   Circle "Kreis_157" at 637,438 size 15x15
      Appearance <- "DB_SDC_ERRORS.EMS[XXX].FC_HOIST_2"
   Circle "Kreis_158" at 637,454 size 15x15
      Appearance <- "DB_SDC_ERRORS.EMS[XXX].FC_HOIST_2"
   Circle "Kreis_159" at 637,470 size 15x15
      Appearance <- "DB_SDC_ERRORS.EMS[XXX].FC_HOIST_2"
   Circle "Kreis_160" at 637,486 size 15x15
      Appearance <- "DB_SDC_ERRORS.EMS[XXX].FC_HOIST_2"
   TextField "Textfeld_248" at 1003,235 size 31x132; Text '501 502 503 504 505 506 507 508 Command forward 501'
   Circle "Kreis_241" at 980,238 size 15x15
      Appearance <- "DB_SDC_ERRORS.EMS[XXX].GEN_1"
   Circle "Kreis_242" at 980,254 size 15x15
      Appearance <- "DB_SDC_ERRORS.EMS[XXX].GEN_1"
   Circle "Kreis_243" at 980,270 size 15x15
      Appearance <- "DB_SDC_ERRORS.EMS[XXX].GEN_1"
   Circle "Kreis_244" at 980,286 size 15x15
      Appearance <- "DB_SDC_ERRORS.EMS[XXX].GEN_1"
   Circle "Kreis_245" at 980,302 size 15x15
      Appearance <- "DB_SDC_ERRORS.EMS[XXX].GEN_1"
   Circle "Kreis_246" at 980,318 size 15x15
      Appearance <- "DB_SDC_ERRORS.EMS[XXX].GEN_1"
   Circle "Kreis_247" at 980,334 size 15x15
      Appearance <- "DB_SDC_ERRORS.EMS[XXX].GEN_1"
   Circle "Kreis_248" at 980,350 size 15x15
      Appearance <- "DB_SDC_ERRORS.EMS[XXX].GEN_1"
   TextField "Textfeld_256" at 1060,235 size 31x132; Text '509 510 511 512 513 514 515 516 Command forward 509'
   Circle "Kreis_249" at 1037,238 size 15x15
      Appearance <- "DB_SDC_ERRORS.EMS[XXX].GEN_1"
   Circle "Kreis_250" at 1037,254 size 15x15
      Appearance <- "DB_SDC_ERRORS.EMS[XXX].GEN_1"
   Circle "Kreis_251" at 1037,270 size 15x15
      Appearance <- "DB_SDC_ERRORS.EMS[XXX].GEN_1"
   Circle "Kreis_252" at 1037,286 size 15x15
      Appearance <- "DB_SDC_ERRORS.EMS[XXX].GEN_1"
   Circle "Kreis_253" at 1037,302 size 15x15
      Appearance <- "DB_SDC_ERRORS.EMS[XXX].GEN_1"
   Circle "Kreis_254" at 1037,318 size 15x15
      Appearance <- "DB_SDC_ERRORS.EMS[XXX].GEN_1"
   Circle "Kreis_255" at 1037,334 size 15x15
      Appearance <- "DB_SDC_ERRORS.EMS[XXX].GEN_1"
   Circle "Kreis_256" at 1037,350 size 15x15
      Appearance <- "DB_SDC_ERRORS.EMS[XXX].GEN_1"
   TextField "Textfeld_264" at 1041,202 size 119x38; Text 'generally / EMS-Number / General'
   Circle "Kreis_257" at 980,374 size 15x15
      Appearance <- "DB_SDC_ERRORS.EMS[XXX].GEN_3"
   Circle "Kreis_258" at 980,390 size 15x15
      Appearance <- "DB_SDC_ERRORS.EMS[XXX].GEN_3"
   Circle "Kreis_259" at 980,406 size 15x15
      Appearance <- "DB_SDC_ERRORS.EMS[XXX].GEN_3"
   Circle "Kreis_260" at 980,422 size 15x15
      Appearance <- "DB_SDC_ERRORS.EMS[XXX].GEN_3"
   Circle "Kreis_261" at 980,438 size 15x15
      Appearance <- "DB_SDC_ERRORS.EMS[XXX].GEN_3"
   Circle "Kreis_262" at 980,454 size 15x15
      Appearance <- "DB_SDC_ERRORS.EMS[XXX].GEN_3"
   Circle "Kreis_263" at 980,470 size 15x15
      Appearance <- "DB_SDC_ERRORS.EMS[XXX].GEN_3"
   Circle "Kreis_264" at 980,486 size 15x15
      Appearance <- "DB_SDC_ERRORS.EMS[XXX].GEN_3"
   Circle "Kreis_265" at 1037,374 size 15x15
      Appearance <- "DB_SDC_ERRORS.EMS[XXX].GEN_3"
   Circle "Kreis_266" at 1037,390 size 15x15
      Appearance <- "DB_SDC_ERRORS.EMS[XXX].GEN_3"
   Circle "Kreis_267" at 1037,406 size 15x15
      Appearance <- "DB_SDC_ERRORS.EMS[XXX].GEN_3"
   Circle "Kreis_268" at 1037,422 size 15x15
      Appearance <- "DB_SDC_ERRORS.EMS[XXX].GEN_3"
   Circle "Kreis_269" at 1037,438 size 15x15
      Appearance <- "DB_SDC_ERRORS.EMS[XXX].GEN_3"
   Circle "Kreis_270" at 1037,454 size 15x15
      Appearance <- "DB_SDC_ERRORS.EMS[XXX].GEN_3"
   Circle "Kreis_271" at 1037,470 size 15x15
      Appearance <- "DB_SDC_ERRORS.EMS[XXX].GEN_3"
   Circle "Kreis_272" at 1037,486 size 15x15
      Appearance <- "DB_SDC_ERRORS.EMS[XXX].GEN_3"
   TextField "Textfeld_281" at 1123,235 size 31x132; Text '517 518 519 520 521 522 523 524 Command forward 517'
   Circle "Kreis_273" at 1100,238 size 15x15
      Appearance <- "DB_SDC_ERRORS.EMS[XXX].GEN_2"
   Circle "Kreis_274" at 1100,254 size 15x15
      Appearance <- "DB_SDC_ERRORS.EMS[XXX].GEN_2"
   Circle "Kreis_275" at 1100,270 size 15x15
      Appearance <- "DB_SDC_ERRORS.EMS[XXX].GEN_2"
   Circle "Kreis_276" at 1100,286 size 15x15
      Appearance <- "DB_SDC_ERRORS.EMS[XXX].GEN_2"
   Circle "Kreis_277" at 1100,302 size 15x15
      Appearance <- "DB_SDC_ERRORS.EMS[XXX].GEN_2"
   Circle "Kreis_278" at 1100,318 size 15x15
      Appearance <- "DB_SDC_ERRORS.EMS[XXX].GEN_2"
   Circle "Kreis_279" at 1100,334 size 15x15
      Appearance <- "DB_SDC_ERRORS.EMS[XXX].GEN_2"
   Circle "Kreis_280" at 1100,350 size 15x15
      Appearance <- "DB_SDC_ERRORS.EMS[XXX].GEN_2"
   TextField "Textfeld_289" at 1180,235 size 31x132; Text '525 526 527 528 529 530 531 532 Command forward 525'
   Circle "Kreis_281" at 1157,238 size 15x15
      Appearance <- "DB_SDC_ERRORS.EMS[XXX].GEN_2"
   Circle "Kreis_282" at 1157,254 size 15x15
      Appearance <- "DB_SDC_ERRORS.EMS[XXX].GEN_2"
   Circle "Kreis_283" at 1157,270 size 15x15
      Appearance <- "DB_SDC_ERRORS.EMS[XXX].GEN_2"
   Circle "Kreis_284" at 1157,286 size 15x15
      Appearance <- "DB_SDC_ERRORS.EMS[XXX].GEN_2"
   Circle "Kreis_285" at 1157,302 size 15x15
      Appearance <- "DB_SDC_ERRORS.EMS[XXX].GEN_2"
   Circle "Kreis_286" at 1157,318 size 15x15
      Appearance <- "DB_SDC_ERRORS.EMS[XXX].GEN_2"
   Circle "Kreis_287" at 1157,334 size 15x15
      Appearance <- "DB_SDC_ERRORS.EMS[XXX].GEN_2"
   Circle "Kreis_288" at 1157,350 size 15x15
      Appearance <- "DB_SDC_ERRORS.EMS[XXX].GEN_2"
   Circle "Kreis_289" at 1100,374 size 15x15
      Appearance <- "DB_SDC_ERRORS.EMS[XXX].GEN_4"
   Circle "Kreis_290" at 1100,390 size 15x15
      Appearance <- "DB_SDC_ERRORS.EMS[XXX].GEN_4"
   Circle "Kreis_291" at 1100,406 size 15x15
      Appearance <- "DB_SDC_ERRORS.EMS[XXX].GEN_4"
   Circle "Kreis_292" at 1100,422 size 15x15
      Appearance <- "DB_SDC_ERRORS.EMS[XXX].GEN_4"
   Circle "Kreis_293" at 1100,438 size 15x15
      Appearance <- "DB_SDC_ERRORS.EMS[XXX].GEN_4"
   Circle "Kreis_294" at 1100,454 size 15x15
      Appearance <- "DB_SDC_ERRORS.EMS[XXX].GEN_4"
   Circle "Kreis_295" at 1100,470 size 15x15
      Appearance <- "DB_SDC_ERRORS.EMS[XXX].GEN_4"
   Circle "Kreis_296" at 1100,486 size 15x15
      Appearance <- "DB_SDC_ERRORS.EMS[XXX].GEN_4"
   Circle "Kreis_297" at 1157,374 size 15x15
      Appearance <- "DB_SDC_ERRORS.EMS[XXX].GEN_4"
   Circle "Kreis_298" at 1157,390 size 15x15
      Appearance <- "DB_SDC_ERRORS.EMS[XXX].GEN_4"
   Circle "Kreis_299" at 1157,406 size 15x15
      Appearance <- "DB_SDC_ERRORS.EMS[XXX].GEN_4"
   Circle "Kreis_300" at 1157,422 size 15x15
      Appearance <- "DB_SDC_ERRORS.EMS[XXX].GEN_4"
   Circle "Kreis_301" at 1157,438 size 15x15
      Appearance <- "DB_SDC_ERRORS.EMS[XXX].GEN_4"
   Circle "Kreis_302" at 1157,454 size 15x15
      Appearance <- "DB_SDC_ERRORS.EMS[XXX].GEN_4"
   Circle "Kreis_303" at 1157,470 size 15x15
      Appearance <- "DB_SDC_ERRORS.EMS[XXX].GEN_4"
   Circle "Kreis_304" at 1157,486 size 15x15
      Appearance <- "DB_SDC_ERRORS.EMS[XXX].GEN_4"
   TextField "Textfeld_313" at 950,250 size 27x114; Text 'errors / EMS-Number / Errors'
   TextField "Textfeld_314" at 950,368 size 27x144; Text 'warnings / EMS-Number / Warnings'
   TextField "Textfeld_265" at 1003,371 size 31x132; Text '801 802 803 804 805 806 807 808 Command forward 801'
   TextField "Textfeld_273" at 1060,371 size 31x132; Text '809 810 811 812 813 814 815 816 Command forward 809'
   TextField "Textfeld_297" at 1123,371 size 31x132; Text '817 818 819 820 821 822 823 824 Command forward 817'
   TextField "Textfeld_305" at 1180,371 size 31x132; Text '825 826 827 828 829 830 831 832 Command forward 825'
   TextField "Textfeld_315" at 1003,531 size 31x132; Text '901 902 903 904 905 906 907 908 Command forward 901'
   Circle "Kreis_305" at 980,534 size 15x15
      Appearance <- "DB_SDC_ERRORS.EMS[XXX].SDC"
   Circle "Kreis_306" at 980,550 size 15x15
      Appearance <- "DB_SDC_ERRORS.EMS[XXX].SDC"
   Circle "Kreis_307" at 980,566 size 15x15
      Appearance <- "DB_SDC_ERRORS.EMS[XXX].SDC"
   Circle "Kreis_308" at 980,582 size 15x15
      Appearance <- "DB_SDC_ERRORS.EMS[XXX].SDC"
   Circle "Kreis_309" at 980,598 size 15x15
      Appearance <- "DB_SDC_ERRORS.EMS[XXX].SDC"
   Circle "Kreis_310" at 980,614 size 15x15
      Appearance <- "DB_SDC_ERRORS.EMS[XXX].SDC"
   Circle "Kreis_311" at 980,630 size 15x15
      Appearance <- "DB_SDC_ERRORS.EMS[XXX].SDC"
   Circle "Kreis_312" at 980,646 size 15x15
      Appearance <- "DB_SDC_ERRORS.EMS[XXX].SDC"
   TextField "Textfeld_323" at 1060,531 size 31x132; Text '909 910 911 912 913 914 915 916 Command forward 909'
   Circle "Kreis_313" at 1037,534 size 15x15
      Appearance <- "DB_SDC_ERRORS.EMS[XXX].SDC"
   Circle "Kreis_314" at 1037,550 size 15x15
      Appearance <- "DB_SDC_ERRORS.EMS[XXX].SDC"
   Circle "Kreis_315" at 1037,566 size 15x15
      Appearance <- "DB_SDC_ERRORS.EMS[XXX].SDC"
   Circle "Kreis_316" at 1037,582 size 15x15
      Appearance <- "DB_SDC_ERRORS.EMS[XXX].SDC"
   Circle "Kreis_317" at 1037,598 size 15x15
      Appearance <- "DB_SDC_ERRORS.EMS[XXX].SDC"
   Circle "Kreis_318" at 1037,614 size 15x15
      Appearance <- "DB_SDC_ERRORS.EMS[XXX].SDC"
   Circle "Kreis_319" at 1037,630 size 15x15
      Appearance <- "DB_SDC_ERRORS.EMS[XXX].SDC"
   Circle "Kreis_320" at 1037,646 size 15x15
      Appearance <- "DB_SDC_ERRORS.EMS[XXX].SDC"
   TextField "Textfeld_331" at 1029,504 size 119x27; Text 'SDC / EMS-Number'
   TextField "Textfeld_348" at 950,566 size 27x61; Text 'EMS / EMS-Number'
   TextField "Textfeld_332" at 953,671 size 27x60; Text 'gen. / EMS-Number / General'
   TextField "Textfeld_333" at 1003,667 size 31x70; Text '917 918 919 920 Command forward 917'
   Circle "Kreis_321" at 980,670 size 15x15
      Appearance <- "DB_SDC_ERRORS.SDC"
   Circle "Kreis_322" at 980,686 size 15x15
      Appearance <- "DB_SDC_ERRORS.SDC"
   Circle "Kreis_323" at 980,702 size 15x15
      Appearance <- "DB_SDC_ERRORS.SDC"
   Circle "Kreis_324" at 980,718 size 15x15
      Appearance <- "DB_SDC_ERRORS.SDC"
   TextField "Textfeld_337" at 1056,667 size 31x70; Text '921 922 923 924 Command forward 921'
   Circle "Kreis_325" at 1037,670 size 15x15
      Appearance <- "DB_SDC_ERRORS.SDC"
   Circle "Kreis_326" at 1037,686 size 15x15
      Appearance <- "DB_SDC_ERRORS.SDC"
   Circle "Kreis_327" at 1037,702 size 15x15
      Appearance <- "DB_SDC_ERRORS.SDC"
   Circle "Kreis_328" at 1037,718 size 15x15
      Appearance <- "DB_SDC_ERRORS.SDC"
   SymbolicIOField "Symbolisches EA-Feld_1" at 592,156 size 626x35; TextOn '1'; TextOff '0'; TextList "SDC_ER_EMS"
      ProcessValue <- "_DB_SDC_ERRORS.Error_nr"
   IOField "EA-Feld_1" at 519,156 size 66x35; FormatPattern 999
      ProcessValue <- "_DB_SDC_ERRORS.Error_nr"
   TextField "Textfeld_341" at 521,129 size 116x27; Text 'ER.Nr. / EMS-Number'
   TextField "Textfeld_342" at 600,129 size 116x27; Text 'ER.Text / EMS-Number'
   Button "Schaltfläche_2" at 207,238 size 59x15; TextOff 'Text'
      on Click: SetTag("_DB_SDC_ERRORS.Error_nr", 601)
   Button "Schaltfläche_4" at 207,254 size 59x15; TextOff 'Text'
      on Click: SetTag("_DB_SDC_ERRORS.Error_nr", 602)
   Button "Schaltfläche_5" at 207,270 size 59x15; TextOff 'Text'
      on Click: SetTag("_DB_SDC_ERRORS.Error_nr", 603)
   Button "Schaltfläche_6" at 207,286 size 59x15; TextOff 'Text'
      on Click: SetTag("_DB_SDC_ERRORS.Error_nr", 604)
   Button "Schaltfläche_7" at 207,302 size 59x15; TextOff 'Text'
      on Click: SetTag("_DB_SDC_ERRORS.Error_nr", 605)
   Button "Schaltfläche_8" at 207,318 size 59x15; TextOff 'Text'
      on Click: SetTag("_DB_SDC_ERRORS.Error_nr", 606)
   Button "Schaltfläche_9" at 207,334 size 59x15; TextOff 'Text'
      on Click: SetTag("_DB_SDC_ERRORS.Error_nr", 607)
   Button "Schaltfläche_10" at 207,350 size 59x15; TextOff 'Text'
      on Click: SetTag("_DB_SDC_ERRORS.Error_nr", 608)
   Button "Schaltfläche_11" at 269,238 size 59x15; TextOff 'Text'
      on Click: SetTag("_DB_SDC_ERRORS.Error_nr", 609)
   Button "Schaltfläche_12" at 269,254 size 59x15; TextOff 'Text'
      on Click: SetTag("_DB_SDC_ERRORS.Error_nr", 610)
   Button "Schaltfläche_13" at 269,270 size 59x15; TextOff 'Text'
      on Click: SetTag("_DB_SDC_ERRORS.Error_nr", 611)
   Button "Schaltfläche_14" at 269,286 size 59x15; TextOff 'Text'
      on Click: SetTag("_DB_SDC_ERRORS.Error_nr", 612)
   Button "Schaltfläche_15" at 269,302 size 59x15; TextOff 'Text'
      on Click: SetTag("_DB_SDC_ERRORS.Error_nr", 613)
   Button "Schaltfläche_16" at 269,318 size 59x15; TextOff 'Text'
      on Click: SetTag("_DB_SDC_ERRORS.Error_nr", 614)
   Button "Schaltfläche_17" at 269,334 size 59x15; TextOff 'Text'
      on Click: SetTag("_DB_SDC_ERRORS.Error_nr", 615)
   Button "Schaltfläche_18" at 269,350 size 59x15; TextOff 'Text'
      on Click: SetTag("_DB_SDC_ERRORS.Error_nr", 616)
   Button "Schaltfläche_19" at 331,238 size 54x15; TextOff 'Text'
      on Click: SetTag("_DB_SDC_ERRORS.Error_nr", 617)
   Button "Schaltfläche_20" at 331,254 size 54x15; TextOff 'Text'
      on Click: SetTag("_DB_SDC_ERRORS.Error_nr", 618)
   Button "Schaltfläche_21" at 331,270 size 54x15; TextOff 'Text'
      on Click: SetTag("_DB_SDC_ERRORS.Error_nr", 619)
   Button "Schaltfläche_22" at 331,286 size 54x15; TextOff 'Text'
      on Click: SetTag("_DB_SDC_ERRORS.Error_nr", 620)
   Button "Schaltfläche_23" at 331,302 size 54x15; TextOff 'Text'
      on Click: SetTag("_DB_SDC_ERRORS.Error_nr", 621)
   Button "Schaltfläche_24" at 331,318 size 54x15; TextOff 'Text'
      on Click: SetTag("_DB_SDC_ERRORS.Error_nr", 622)
   Button "Schaltfläche_25" at 331,334 size 54x15; TextOff 'Text'
      on Click: SetTag("_DB_SDC_ERRORS.Error_nr", 623)
   Button "Schaltfläche_26" at 331,350 size 54x15; TextOff 'Text'
      on Click: SetTag("_DB_SDC_ERRORS.Error_nr", 624)
   Button "Schaltfläche_27" at 388,238 size 59x15; TextOff 'Text'
      on Click: SetTag("_DB_SDC_ERRORS.Error_nr", 625)
   Button "Schaltfläche_28" at 388,254 size 59x15; TextOff 'Text'
      on Click: SetTag("_DB_SDC_ERRORS.Error_nr", 626)
   Button "Schaltfläche_29" at 388,270 size 59x15; TextOff 'Text'
      on Click: SetTag("_DB_SDC_ERRORS.Error_nr", 627)
   Button "Schaltfläche_30" at 388,286 size 59x15; TextOff 'Text'
      on Click: SetTag("_DB_SDC_ERRORS.Error_nr", 628)
   Button "Schaltfläche_31" at 388,302 size 59x15; TextOff 'Text'
      on Click: SetTag("_DB_SDC_ERRORS.Error_nr", 629)
   Button "Schaltfläche_32" at 388,318 size 59x15; TextOff 'Text'
      on Click: SetTag("_DB_SDC_ERRORS.Error_nr", 630)
   Button "Schaltfläche_33" at 388,334 size 59x15; TextOff 'Text'
      on Click: SetTag("_DB_SDC_ERRORS.Error_nr", 631)
   Button "Schaltfläche_34" at 388,350 size 59x15; TextOff 'Text'
      on Click: SetTag("_DB_SDC_ERRORS.Error_nr", 632)
   Button "Schaltfläche_35" at 206,374 size 59x15; TextOff 'Text'
      on Click: SetTag("_DB_SDC_ERRORS.Error_nr", 633)
   Button "Schaltfläche_36" at 206,390 size 59x15; TextOff 'Text'
      on Click: SetTag("_DB_SDC_ERRORS.Error_nr", 634)
   Button "Schaltfläche_37" at 206,406 size 59x15; TextOff 'Text'
      on Click: SetTag("_DB_SDC_ERRORS.Error_nr", 635)
   Button "Schaltfläche_38" at 206,422 size 59x15; TextOff 'Text'
      on Click: SetTag("_DB_SDC_ERRORS.Error_nr", 636)
   Button "Schaltfläche_39" at 206,438 size 59x15; TextOff 'Text'
      on Click: SetTag("_DB_SDC_ERRORS.Error_nr", 637)
   Button "Schaltfläche_40" at 206,454 size 59x15; TextOff 'Text'
      on Click: SetTag("_DB_SDC_ERRORS.Error_nr", 638)
   Button "Schaltfläche_41" at 206,470 size 59x15; TextOff 'Text'
      on Click: SetTag("_DB_SDC_ERRORS.Error_nr", 639)
   Button "Schaltfläche_42" at 206,486 size 59x15; TextOff 'Text'
      on Click: SetTag("_DB_SDC_ERRORS.Error_nr", 640)
   Button "Schaltfläche_43" at 268,374 size 59x15; TextOff 'Text'
      on Click: SetTag("_DB_SDC_ERRORS.Error_nr", 641)
   Button "Schaltfläche_44" at 268,390 size 59x15; TextOff 'Text'
      on Click: SetTag("_DB_SDC_ERRORS.Error_nr", 642)
   Button "Schaltfläche_45" at 268,406 size 59x15; TextOff 'Text'
      on Click: SetTag("_DB_SDC_ERRORS.Error_nr", 643)
   Button "Schaltfläche_46" at 268,422 size 59x15; TextOff 'Text'
      on Click: SetTag("_DB_SDC_ERRORS.Error_nr", 644)
   Button "Schaltfläche_47" at 268,438 size 59x15; TextOff 'Text'
      on Click: SetTag("_DB_SDC_ERRORS.Error_nr", 645)
   Button "Schaltfläche_48" at 268,454 size 59x15; TextOff 'Text'
      on Click: SetTag("_DB_SDC_ERRORS.Error_nr", 646)
   Button "Schaltfläche_49" at 268,470 size 59x15; TextOff 'Text'
      on Click: SetTag("_DB_SDC_ERRORS.Error_nr", 647)
   Button "Schaltfläche_50" at 268,486 size 59x15; TextOff 'Text'
      on Click: SetTag("_DB_SDC_ERRORS.Error_nr", 648)
   Button "Schaltfläche_51" at 207,510 size 59x15; TextOff 'Text'
      on Click: SetTag("_DB_SDC_ERRORS.Error_nr", 649)
   Button "Schaltfläche_52" at 207,526 size 59x15; TextOff 'Text'
      on Click: SetTag("_DB_SDC_ERRORS.Error_nr", 650)
   Button "Schaltfläche_53" at 207,542 size 59x15; TextOff 'Text'
      on Click: SetTag("_DB_SDC_ERRORS.Error_nr", 651)
   Button "Schaltfläche_54" at 207,558 size 59x15; TextOff 'Text'
      on Click: SetTag("_DB_SDC_ERRORS.Error_nr", 652)
   Button "Schaltfläche_55" at 207,574 size 59x15; TextOff 'Text'
      on Click: SetTag("_DB_SDC_ERRORS.Error_nr", 653)
   Button "Schaltfläche_56" at 207,590 size 59x15; TextOff 'Text'
      on Click: SetTag("_DB_SDC_ERRORS.Error_nr", 654)
   Button "Schaltfläche_57" at 207,606 size 59x15; TextOff 'Text'
      on Click: SetTag("_DB_SDC_ERRORS.Error_nr", 655)
   Button "Schaltfläche_58" at 207,622 size 59x15; TextOff 'Text'
      on Click: SetTag("_DB_SDC_ERRORS.Error_nr", 656)
   Button "Schaltfläche_59" at 269,510 size 59x15; TextOff 'Text'
      on Click: SetTag("_DB_SDC_ERRORS.Error_nr", 657)
   Button "Schaltfläche_60" at 269,526 size 59x15; TextOff 'Text'
      on Click: SetTag("_DB_SDC_ERRORS.Error_nr", 658)
   Button "Schaltfläche_61" at 269,542 size 59x15; TextOff 'Text'
      on Click: SetTag("_DB_SDC_ERRORS.Error_nr", 659)
   Button "Schaltfläche_62" at 269,558 size 59x15; TextOff 'Text'
      on Click: SetTag("_DB_SDC_ERRORS.Error_nr", 660)
   Button "Schaltfläche_63" at 269,574 size 59x15; TextOff 'Text'
      on Click: SetTag("_DB_SDC_ERRORS.Error_nr", 661)
   Button "Schaltfläche_64" at 269,590 size 59x15; TextOff 'Text'
      on Click: SetTag("_DB_SDC_ERRORS.Error_nr", 662)
   Button "Schaltfläche_65" at 269,606 size 59x15; TextOff 'Text'
      on Click: SetTag("_DB_SDC_ERRORS.Error_nr", 663)
   Button "Schaltfläche_66" at 269,622 size 59x15; TextOff 'Text'
      on Click: SetTag("_DB_SDC_ERRORS.Error_nr", 664)
   Button "Schaltfläche_67" at 453,237 size 59x15; TextOff 'Text'
      on Click: SetTag("_DB_SDC_ERRORS.Error_nr", 701)
   Button "Schaltfläche_68" at 453,253 size 59x15; TextOff 'Text'
      on Click: SetTag("_DB_SDC_ERRORS.Error_nr", 702)
   Button "Schaltfläche_69" at 453,269 size 59x15; TextOff 'Text'
      on Click: SetTag("_DB_SDC_ERRORS.Error_nr", 703)
   Button "Schaltfläche_70" at 453,285 size 59x15; TextOff 'Text'
      on Click: SetTag("_DB_SDC_ERRORS.Error_nr", 704)
   Button "Schaltfläche_71" at 453,301 size 59x15; TextOff 'Text'
      on Click: SetTag("_DB_SDC_ERRORS.Error_nr", 705)
   Button "Schaltfläche_72" at 453,317 size 59x15; TextOff 'Text'
      on Click: SetTag("_DB_SDC_ERRORS.Error_nr", 706)
   Button "Schaltfläche_73" at 453,333 size 59x15; TextOff 'Text'
      on Click: SetTag("_DB_SDC_ERRORS.Error_nr", 707)
   Button "Schaltfläche_74" at 453,349 size 59x15; TextOff 'Text'
      on Click: SetTag("_DB_SDC_ERRORS.Error_nr", 708)
   Button "Schaltfläche_75" at 515,237 size 59x15; TextOff 'Text'
      on Click: SetTag("_DB_SDC_ERRORS.Error_nr", 709)
   Button "Schaltfläche_76" at 515,253 size 59x15; TextOff 'Text'
      on Click: SetTag("_DB_SDC_ERRORS.Error_nr", 710)
   Button "Schaltfläche_77" at 515,269 size 59x15; TextOff 'Text'
      on Click: SetTag("_DB_SDC_ERRORS.Error_nr", 711)
   Button "Schaltfläche_78" at 515,285 size 59x15; TextOff 'Text'
      on Click: SetTag("_DB_SDC_ERRORS.Error_nr", 712)
   Button "Schaltfläche_79" at 515,301 size 59x15; TextOff 'Text'
      on Click: SetTag("_DB_SDC_ERRORS.Error_nr", 713)
   Button "Schaltfläche_80" at 515,317 size 59x15; TextOff 'Text'
      on Click: SetTag("_DB_SDC_ERRORS.Error_nr", 714)
   Button "Schaltfläche_81" at 515,333 size 59x15; TextOff 'Text'
      on Click: SetTag("_DB_SDC_ERRORS.Error_nr", 715)
   Button "Schaltfläche_82" at 515,349 size 59x15; TextOff 'Text'
      on Click: SetTag("_DB_SDC_ERRORS.Error_nr", 716)
   Button "Schaltfläche_83" at 577,237 size 54x15; TextOff 'Text'
      on Click: SetTag("_DB_SDC_ERRORS.Error_nr", 717)
   Button "Schaltfläche_84" at 577,253 size 54x15; TextOff 'Text'
      on Click: SetTag("_DB_SDC_ERRORS.Error_nr", 718)
   Button "Schaltfläche_85" at 577,269 size 54x15; TextOff 'Text'
      on Click: SetTag("_DB_SDC_ERRORS.Error_nr", 719)
   Button "Schaltfläche_86" at 577,285 size 54x15; TextOff 'Text'
      on Click: SetTag("_DB_SDC_ERRORS.Error_nr", 720)
   Button "Schaltfläche_87" at 577,301 size 54x15; TextOff 'Text'
      on Click: SetTag("_DB_SDC_ERRORS.Error_nr", 721)
   Button "Schaltfläche_88" at 577,317 size 54x15; TextOff 'Text'
      on Click: SetTag("_DB_SDC_ERRORS.Error_nr", 722)
   Button "Schaltfläche_89" at 577,333 size 54x15; TextOff 'Text'
      on Click: SetTag("_DB_SDC_ERRORS.Error_nr", 723)
   Button "Schaltfläche_90" at 577,349 size 54x15; TextOff 'Text'
      on Click: SetTag("_DB_SDC_ERRORS.Error_nr", 724)
   Button "Schaltfläche_91" at 634,237 size 59x15; TextOff 'Text'
      on Click: SetTag("_DB_SDC_ERRORS.Error_nr", 725)
   Button "Schaltfläche_92" at 634,253 size 59x15; TextOff 'Text'
      on Click: SetTag("_DB_SDC_ERRORS.Error_nr", 726)
   Button "Schaltfläche_93" at 634,269 size 59x15; TextOff 'Text'
      on Click: SetTag("_DB_SDC_ERRORS.Error_nr", 727)
   Button "Schaltfläche_94" at 634,285 size 59x15; TextOff 'Text'
      on Click: SetTag("_DB_SDC_ERRORS.Error_nr", 728)
   Button "Schaltfläche_95" at 634,301 size 59x15; TextOff 'Text'
      on Click: SetTag("_DB_SDC_ERRORS.Error_nr", 729)
   Button "Schaltfläche_96" at 634,317 size 59x15; TextOff 'Text'
      on Click: SetTag("_DB_SDC_ERRORS.Error_nr", 730)
   Button "Schaltfläche_97" at 634,333 size 59x15; TextOff 'Text'
      on Click: SetTag("_DB_SDC_ERRORS.Error_nr", 731)
   Button "Schaltfläche_98" at 634,349 size 59x15; TextOff 'Text'
      on Click: SetTag("_DB_SDC_ERRORS.Error_nr", 732)
   Button "Schaltfläche_99" at 452,373 size 59x15; TextOff 'Text'
      on Click: SetTag("_DB_SDC_ERRORS.Error_nr", 733)
   Button "Schaltfläche_100" at 452,389 size 59x15; TextOff 'Text'
      on Click: SetTag("_DB_SDC_ERRORS.Error_nr", 734)
   Button "Schaltfläche_101" at 452,405 size 59x15; TextOff 'Text'
      on Click: SetTag("_DB_SDC_ERRORS.Error_nr", 735)
   Button "Schaltfläche_102" at 452,421 size 59x15; TextOff 'Text'
      on Click: SetTag("_DB_SDC_ERRORS.Error_nr", 736)
   Button "Schaltfläche_103" at 452,437 size 59x15; TextOff 'Text'
      on Click: SetTag("_DB_SDC_ERRORS.Error_nr", 737)
   Button "Schaltfläche_104" at 452,453 size 59x15; TextOff 'Text'
      on Click: SetTag("_DB_SDC_ERRORS.Error_nr", 738)
   Button "Schaltfläche_105" at 452,469 size 59x15; TextOff 'Text'
      on Click: SetTag("_DB_SDC_ERRORS.Error_nr", 739)
   Button "Schaltfläche_106" at 452,485 size 59x15; TextOff 'Text'
      on Click: SetTag("_DB_SDC_ERRORS.Error_nr", 740)
   Button "Schaltfläche_107" at 514,373 size 59x15; TextOff 'Text'
      on Click: SetTag("_DB_SDC_ERRORS.Error_nr", 741)
   Button "Schaltfläche_108" at 514,389 size 59x15; TextOff 'Text'
      on Click: SetTag("_DB_SDC_ERRORS.Error_nr", 742)
   Button "Schaltfläche_109" at 514,405 size 59x15; TextOff 'Text'
      on Click: SetTag("_DB_SDC_ERRORS.Error_nr", 743)
   Button "Schaltfläche_110" at 514,421 size 59x15; TextOff 'Text'
      on Click: SetTag("_DB_SDC_ERRORS.Error_nr", 744)
   Button "Schaltfläche_111" at 514,437 size 59x15; TextOff 'Text'
      on Click: SetTag("_DB_SDC_ERRORS.Error_nr", 745)
   Button "Schaltfläche_112" at 514,453 size 59x15; TextOff 'Text'
      on Click: SetTag("_DB_SDC_ERRORS.Error_nr", 746)
   Button "Schaltfläche_113" at 514,469 size 59x15; TextOff 'Text'
      on Click: SetTag("_DB_SDC_ERRORS.Error_nr", 747)
   Button "Schaltfläche_114" at 514,485 size 59x15; TextOff 'Text'
      on Click: SetTag("_DB_SDC_ERRORS.Error_nr", 748)
   Button "Schaltfläche_115" at 453,509 size 59x15; TextOff 'Text'
      on Click: SetTag("_DB_SDC_ERRORS.Error_nr", 749)
   Button "Schaltfläche_116" at 453,525 size 59x15; TextOff 'Text'
      on Click: SetTag("_DB_SDC_ERRORS.Error_nr", 750)
   Button "Schaltfläche_117" at 453,541 size 59x15; TextOff 'Text'
      on Click: SetTag("_DB_SDC_ERRORS.Error_nr", 751)
   Button "Schaltfläche_118" at 453,557 size 59x15; TextOff 'Text'
      on Click: SetTag("_DB_SDC_ERRORS.Error_nr", 752)
   Button "Schaltfläche_119" at 453,573 size 59x15; TextOff 'Text'
      on Click: SetTag("_DB_SDC_ERRORS.Error_nr", 753)
   Button "Schaltfläche_120" at 453,589 size 59x15; TextOff 'Text'
      on Click: SetTag("_DB_SDC_ERRORS.Error_nr", 754)
   Button "Schaltfläche_121" at 453,605 size 59x15; TextOff 'Text'
      on Click: SetTag("_DB_SDC_ERRORS.Error_nr", 755)
   Button "Schaltfläche_122" at 453,621 size 59x15; TextOff 'Text'
      on Click: SetTag("_DB_SDC_ERRORS.Error_nr", 756)
   Button "Schaltfläche_123" at 515,509 size 59x15; TextOff 'Text'
      on Click: SetTag("_DB_SDC_ERRORS.Error_nr", 757)
   Button "Schaltfläche_124" at 515,525 size 59x15; TextOff 'Text'
      on Click: SetTag("_DB_SDC_ERRORS.Error_nr", 758)
   Button "Schaltfläche_125" at 515,541 size 59x15; TextOff 'Text'
      on Click: SetTag("_DB_SDC_ERRORS.Error_nr", 759)
   Button "Schaltfläche_126" at 515,557 size 59x15; TextOff 'Text'
      on Click: SetTag("_DB_SDC_ERRORS.Error_nr", 760)
   Button "Schaltfläche_127" at 515,573 size 59x15; TextOff 'Text'
      on Click: SetTag("_DB_SDC_ERRORS.Error_nr", 761)
   Button "Schaltfläche_128" at 515,589 size 59x15; TextOff 'Text'
      on Click: SetTag("_DB_SDC_ERRORS.Error_nr", 762)
   Button "Schaltfläche_129" at 515,605 size 59x15; TextOff 'Text'
      on Click: SetTag("_DB_SDC_ERRORS.Error_nr", 763)
   Button "Schaltfläche_130" at 515,621 size 59x15; TextOff 'Text'
      on Click: SetTag("_DB_SDC_ERRORS.Error_nr", 764)
   Button "Schaltfläche_195" at 973,237 size 59x15; TextOff 'Text'
      on Click: SetTag("_DB_SDC_ERRORS.Error_nr", 501)
   Button "Schaltfläche_196" at 973,253 size 59x15; TextOff 'Text'
      on Click: SetTag("_DB_SDC_ERRORS.Error_nr", 502)
   Button "Schaltfläche_197" at 973,269 size 59x15; TextOff 'Text'
      on Click: SetTag("_DB_SDC_ERRORS.Error_nr", 503)
   Button "Schaltfläche_198" at 973,285 size 59x15; TextOff 'Text'
      on Click: SetTag("_DB_SDC_ERRORS.Error_nr", 504)
   Button "Schaltfläche_199" at 973,301 size 59x15; TextOff 'Text'
      on Click: SetTag("_DB_SDC_ERRORS.Error_nr", 505)
   Button "Schaltfläche_200" at 973,317 size 59x15; TextOff 'Text'
      on Click: SetTag("_DB_SDC_ERRORS.Error_nr", 506)
   Button "Schaltfläche_201" at 973,333 size 59x15; TextOff 'Text'
      on Click: SetTag("_DB_SDC_ERRORS.Error_nr", 507)
   Button "Schaltfläche_202" at 973,349 size 59x15; TextOff 'Text'
      on Click: SetTag("_DB_SDC_ERRORS.Error_nr", 508)
   Button "Schaltfläche_203" at 1035,237 size 59x15; TextOff 'Text'
      on Click: SetTag("_DB_SDC_ERRORS.Error_nr", 509)
   Button "Schaltfläche_204" at 1035,253 size 59x15; TextOff 'Text'
      on Click: SetTag("_DB_SDC_ERRORS.Error_nr", 510)
   Button "Schaltfläche_205" at 1035,269 size 59x15; TextOff 'Text'
      on Click: SetTag("_DB_SDC_ERRORS.Error_nr", 511)
   Button "Schaltfläche_206" at 1035,285 size 59x15; TextOff 'Text'
      on Click: SetTag("_DB_SDC_ERRORS.Error_nr", 512)
   Button "Schaltfläche_207" at 1035,301 size 59x15; TextOff 'Text'
      on Click: SetTag("_DB_SDC_ERRORS.Error_nr", 513)
   Button "Schaltfläche_208" at 1035,317 size 59x15; TextOff 'Text'
      on Click: SetTag("_DB_SDC_ERRORS.Error_nr", 514)
   Button "Schaltfläche_209" at 1035,333 size 59x15; TextOff 'Text'
      on Click: SetTag("_DB_SDC_ERRORS.Error_nr", 515)
   Button "Schaltfläche_210" at 1035,349 size 59x15; TextOff 'Text'
      on Click: SetTag("_DB_SDC_ERRORS.Error_nr", 516)
   Button "Schaltfläche_211" at 1097,237 size 54x15; TextOff 'Text'
      on Click: SetTag("_DB_SDC_ERRORS.Error_nr", 517)
   Button "Schaltfläche_212" at 1097,253 size 54x15; TextOff 'Text'
      on Click: SetTag("_DB_SDC_ERRORS.Error_nr", 518)
   Button "Schaltfläche_213" at 1097,269 size 54x15; TextOff 'Text'
      on Click: SetTag("_DB_SDC_ERRORS.Error_nr", 519)
   Button "Schaltfläche_214" at 1097,285 size 54x15; TextOff 'Text'
      on Click: SetTag("_DB_SDC_ERRORS.Error_nr", 520)
   Button "Schaltfläche_215" at 1097,301 size 54x15; TextOff 'Text'
      on Click: SetTag("_DB_SDC_ERRORS.Error_nr", 521)
   Button "Schaltfläche_216" at 1097,317 size 54x15; TextOff 'Text'
      on Click: SetTag("_DB_SDC_ERRORS.Error_nr", 522)
   Button "Schaltfläche_217" at 1097,333 size 54x15; TextOff 'Text'
      on Click: SetTag("_DB_SDC_ERRORS.Error_nr", 523)
   Button "Schaltfläche_218" at 1097,349 size 54x15; TextOff 'Text'
      on Click: SetTag("_DB_SDC_ERRORS.Error_nr", 524)
   Button "Schaltfläche_219" at 1154,237 size 59x15; TextOff 'Text'
      on Click: SetTag("_DB_SDC_ERRORS.Error_nr", 525)
   Button "Schaltfläche_220" at 1154,253 size 59x15; TextOff 'Text'
      on Click: SetTag("_DB_SDC_ERRORS.Error_nr", 526)
   Button "Schaltfläche_221" at 1154,269 size 59x15; TextOff 'Text'
      on Click: SetTag("_DB_SDC_ERRORS.Error_nr", 527)
   Button "Schaltfläche_222" at 1154,285 size 59x15; TextOff 'Text'
      on Click: SetTag("_DB_SDC_ERRORS.Error_nr", 528)
   Button "Schaltfläche_223" at 1154,301 size 59x15; TextOff 'Text'
      on Click: SetTag("_DB_SDC_ERRORS.Error_nr", 529)
   Button "Schaltfläche_224" at 1154,317 size 59x15; TextOff 'Text'
      on Click: SetTag("_DB_SDC_ERRORS.Error_nr", 530)
   Button "Schaltfläche_225" at 1154,333 size 59x15; TextOff 'Text'
      on Click: SetTag("_DB_SDC_ERRORS.Error_nr", 531)
   Button "Schaltfläche_226" at 1154,349 size 59x15; TextOff 'Text'
      on Click: SetTag("_DB_SDC_ERRORS.Error_nr", 532)
   Button "Schaltfläche_227" at 973,373 size 59x15; TextOff 'Text'
      on Click: SetTag("_DB_SDC_ERRORS.Error_nr", 801)
   Button "Schaltfläche_228" at 973,389 size 59x15; TextOff 'Text'
      on Click: SetTag("_DB_SDC_ERRORS.Error_nr", 802)
   Button "Schaltfläche_229" at 973,405 size 59x15; TextOff 'Text'
      on Click: SetTag("_DB_SDC_ERRORS.Error_nr", 803)
   Button "Schaltfläche_230" at 973,421 size 59x15; TextOff 'Text'
      on Click: SetTag("_DB_SDC_ERRORS.Error_nr", 804)
   Button "Schaltfläche_231" at 973,437 size 59x15; TextOff 'Text'
      on Click: SetTag("_DB_SDC_ERRORS.Error_nr", 805)
   Button "Schaltfläche_232" at 973,453 size 59x15; TextOff 'Text'
      on Click: SetTag("_DB_SDC_ERRORS.Error_nr", 806)
   Button "Schaltfläche_233" at 973,469 size 59x15; TextOff 'Text'
      on Click: SetTag("_DB_SDC_ERRORS.Error_nr", 807)
   Button "Schaltfläche_234" at 973,485 size 59x15; TextOff 'Text'
      on Click: SetTag("_DB_SDC_ERRORS.Error_nr", 808)
   Button "Schaltfläche_235" at 1035,373 size 59x15; TextOff 'Text'
      on Click: SetTag("_DB_SDC_ERRORS.Error_nr", 809)
   Button "Schaltfläche_236" at 1035,389 size 59x15; TextOff 'Text'
      on Click: SetTag("_DB_SDC_ERRORS.Error_nr", 810)
   Button "Schaltfläche_237" at 1035,405 size 59x15; TextOff 'Text'
      on Click: SetTag("_DB_SDC_ERRORS.Error_nr", 811)
   Button "Schaltfläche_238" at 1035,421 size 59x15; TextOff 'Text'
      on Click: SetTag("_DB_SDC_ERRORS.Error_nr", 812)
   Button "Schaltfläche_239" at 1035,437 size 59x15; TextOff 'Text'
      on Click: SetTag("_DB_SDC_ERRORS.Error_nr", 813)
   Button "Schaltfläche_240" at 1035,453 size 59x15; TextOff 'Text'
      on Click: SetTag("_DB_SDC_ERRORS.Error_nr", 814)
   Button "Schaltfläche_241" at 1035,469 size 59x15; TextOff 'Text'
      on Click: SetTag("_DB_SDC_ERRORS.Error_nr", 815)
   Button "Schaltfläche_242" at 1035,485 size 59x15; TextOff 'Text'
      on Click: SetTag("_DB_SDC_ERRORS.Error_nr", 816)
   Button "Schaltfläche_243" at 1097,373 size 54x15; TextOff 'Text'
      on Click: SetTag("_DB_SDC_ERRORS.Error_nr", 817)
   Button "Schaltfläche_244" at 1097,389 size 54x15; TextOff 'Text'
      on Click: SetTag("_DB_SDC_ERRORS.Error_nr", 818)
   Button "Schaltfläche_245" at 1097,405 size 54x15; TextOff 'Text'
      on Click: SetTag("_DB_SDC_ERRORS.Error_nr", 819)
   Button "Schaltfläche_246" at 1097,421 size 54x15; TextOff 'Text'
      on Click: SetTag("_DB_SDC_ERRORS.Error_nr", 820)
   Button "Schaltfläche_247" at 1097,437 size 54x15; TextOff 'Text'
      on Click: SetTag("_DB_SDC_ERRORS.Error_nr", 821)
   Button "Schaltfläche_248" at 1097,453 size 54x15; TextOff 'Text'
      on Click: SetTag("_DB_SDC_ERRORS.Error_nr", 822)
   Button "Schaltfläche_249" at 1097,469 size 54x15; TextOff 'Text'
      on Click: SetTag("_DB_SDC_ERRORS.Error_nr", 823)
   Button "Schaltfläche_250" at 1097,485 size 54x15; TextOff 'Text'
      on Click: SetTag("_DB_SDC_ERRORS.Error_nr", 824)
   Button "Schaltfläche_251" at 1154,373 size 59x15; TextOff 'Text'
      on Click: SetTag("_DB_SDC_ERRORS.Error_nr", 825)
   Button "Schaltfläche_252" at 1154,389 size 59x15; TextOff 'Text'
      on Click: SetTag("_DB_SDC_ERRORS.Error_nr", 826)
   Button "Schaltfläche_253" at 1154,405 size 59x15; TextOff 'Text'
      on Click: SetTag("_DB_SDC_ERRORS.Error_nr", 827)
   Button "Schaltfläche_254" at 1154,421 size 59x15; TextOff 'Text'
      on Click: SetTag("_DB_SDC_ERRORS.Error_nr", 828)
   Button "Schaltfläche_255" at 1154,437 size 59x15; TextOff 'Text'
      on Click: SetTag("_DB_SDC_ERRORS.Error_nr", 829)
